// TIA Portal project "Delta_Praktika_P&P" (V17) (continued)

               // jog to position
               //*********************************************************************************************************
             ELSIF #tempJogToPosition THEN
               // set jog target position and configuration
               #instMC_MoveLinearAbsoute.Position[1] := #targetPosition.x;
               #instMC_MoveLinearAbsoute.Position[2] := #targetPosition.y;
               #instMC_MoveLinearAbsoute.Position[3] := #targetPosition.z;
               #instMC_MoveLinearAbsoute.Position[4] := #targetPosition.a;
               #instMC_MoveLinearAbsoute.CoordSystem := #coordSystem;
               #instMC_MoveLinearAbsoute.Velocity := #dynamics.path.velocity;
               #instMC_MoveLinearAbsoute.Acceleration := #dynamics.path.acceleration;
               #instMC_MoveLinearAbsoute.Deceleration := #dynamics.path.deceleration;
               #instMC_MoveLinearAbsoute.Jerk := #dynamics.path.jerk;
               #instMC_MoveLinearAbsoute.DynamicAdaption := #dynamics.dynamicAdaption;
               #instMC_MoveLinearAbsoute.DirectionA := #dynamics.directionA;

               // jog synchronous point to point
               //*********************************************************************************************************
             ELSIF #tempJogSPTP THEN
               #instMC_MoveDirectAbsolute.Position[1] := #targetPosition.x;
               #instMC_MoveDirectAbsolute.Position[2] := #targetPosition.y;
               #instMC_MoveDirectAbsolute.Position[3] := #targetPosition.z;
               #instMC_MoveDirectAbsolute.Position[4] := #targetPosition.a;
               #instMC_MoveDirectAbsolute.CoordSystem := #coordSystem;
               #instMC_MoveDirectAbsolute.VelocityFactor := #dynamics.sPTP.velocityFactor;
               #instMC_MoveDirectAbsolute.AccelerationFactor := #dynamics.sPTP.accelerationFactor;
               #instMC_MoveDirectAbsolute.DecelerationFactor := #dynamics.sPTP.decelerationFactor;
               #instMC_MoveDirectAbsolute.JerkFactor := #dynamics.sPTP.jerkFactor;
               #instMC_MoveDirectAbsolute.LinkConstellation := #linkconstellation;
               #instMC_MoveDirectAbsolute.PositionMode := 1;
               #instMC_MoveDirectAbsolute.DirectionA := #dynamics.directionA;

             END_IF;

           END_REGION

           REGION SET_ORIENTATION_DYNAMICS

             IF (((#jogDirection = 4) AND (#tempJogForward OR #tempJogBackward)) OR #tempJogToPosition)
               AND (#dynamics.orientation.velocity > 0.0 // check if change of orientation dynamics is required
               OR #dynamics.orientation.acceleration > 0.0
               OR #dynamics.orientation.deceleration > 0.0
               OR #dynamics.orientation.jerk > 0.0)
             THEN
               // safe default dynamics for orientation axis
               #statOrientationDynamicsOld.velocity := #axesGroup.DynamicDefaults.Orientation.Velocity;
               #statOrientationDynamicsOld.acceleration := #axesGroup.DynamicDefaults.Orientation.Acceleration;
               #statOrientationDynamicsOld.deceleration := #axesGroup.DynamicDefaults.Orientation.Deceleration;
               #statOrientationDynamicsOld.jerk := #axesGroup.DynamicDefaults.Orientation.Jerk;

               // change orientation default dynamics temporary
               IF #dynamics.orientation.velocity > 0.0 THEN
                 #axesGroup.DynamicDefaults.Orientation.Velocity := #dynamics.orientation.velocity;
               END_IF;
               IF #dynamics.orientation.acceleration > 0.0 THEN
                 #axesGroup.DynamicDefaults.Orientation.Acceleration := #dynamics.orientation.acceleration;
               END_IF;
               IF #dynamics.orientation.deceleration > 0.0 THEN
                 #axesGroup.DynamicDefaults.Orientation.Deceleration := #dynamics.orientation.deceleration;
               END_IF;
               IF #dynamics.orientation.jerk > 0.0 THEN
                 #axesGroup.DynamicDefaults.Orientation.Jerk := #dynamics.orientation.jerk;
               END_IF;

               // Orientation default dynamics will be reseted to previous values after jogging
               #statOrientationDynamicsChanged := TRUE;
             END_IF;
           END_REGION

           REGION STATE_TRANSITION

             // check if change of tool is required
             IF (#tool <> #statToolOld) THEN
               #statFBState := #FB_STATE_SET_TOOL;
             ELSE // execute movement
               #statFBState := #FB_STATE_EXECUTE_MOVEMENT;
             END_IF;

           END_REGION

         END_IF;

       #FB_STATE_SET_TOOL:

         REGION TOOL_CHANGE

           IF #axesGroup.StatusWord.%X6 // no motion command is acitve
             AND NOT #axesGroup.StatusWord.%X17 // not interrupted
             AND #axesGroup.StatusWord.%X12 // constant velocity
           THEN
             #instMC_SetTool.Execute := TRUE;
             #instMC_SetTool.ToolNumber := #tool;
           END_IF;

         END_REGION

         REGION STATE_TRANSITION

           // tool has been changed
           IF #instMC_SetTool.Done THEN
             #statToolOld := #tool;
             #statFBState := #FB_STATE_EXECUTE_MOVEMENT;
           END_IF;

         END_REGION

       #FB_STATE_EXECUTE_MOVEMENT:

         REGION SET_JOG_COMMAND

             // Cartesian jogging
             IF (#tempJogForward OR #tempJogBackward) THEN
               #instMC_MoveLinearRelative.Execute := TRUE;

               // jog to target position  
             ELSIF #tempJogToPosition THEN
               #instMC_MoveLinearAbsoute.Execute := TRUE;

               //jog synchronous point to point
             ELSIF #tempJogSPTP THEN
               #instMC_MoveDirectAbsolute.Execute := TRUE;

             ELSE
               #instMC_MoveLinearRelative.Execute := FALSE;
               #instMC_MoveLinearAbsoute.Execute := FALSE;
               #instMC_MoveDirectAbsolute.Execute := FALSE;
             END_IF;

         END_REGION

         REGION STATE_TRANSITION

           IF #instMC_MoveLinearRelative.Done OR #instMC_MoveLinearAbsoute.Done OR #instMC_MoveDirectAbsolute.Done THEN
             #statStatus := #STATUS_EXECUTION_FINISHED;
           END_IF;

         END_REGION

       #FB_STATE_STOP:

         REGION STOP_KINEMATICS_MOTION

           // set execute if group stop not busy
           #instMC_GroupStop.Execute := (NOT #instMC_GroupStop.Busy AND NOT #instMC_GroupStop.Done AND NOT #instMC_GroupStop.Error);

         END_REGION

         REGION STATE_TRANSITION

           IF (#instMC_GroupStop.Done AND #axesGroup.StatusWord.%X6) THEN // Added X6 according to AW
             #statStatus := #STATUS_EXECUTION_FINISHED;
           ELSIF #axesGroup.StatusWord.%X1 THEN // general TO error
             #statStatus := #ERR_TO_KINEMATICS;
           ELSIF #instMC_MoveLinearRelative.Error THEN
             #statStatus := #instMC_MoveLinearRelative.ErrorId;
           ELSIF #instMC_MoveLinearAbsoute.Error THEN
             #statStatus := #instMC_MoveLinearAbsoute.ErrorId;
           ELSIF #instMC_MoveDirectAbsolute.Error THEN
             #statStatus := #instMC_MoveDirectAbsolute.ErrorId;
           ELSIF #instMC_SetTool.Error THEN
             #statStatus := #instMC_SetTool.ErrorId;
           ELSIF #instMC_GroupStop.Error THEN
             #statStatus := #instMC_GroupStop.ErrorId;
           END_IF;

         END_REGION

       ELSE // Undefined state in state machine reached
         #statStatus := #ERR_UNDEFINED_STATE;
     END_CASE;

   END_REGION STATE_MACHINE

   REGION OUTPUTS

     // Write outputs
     IF (#statStatus = #STATUS_EXECUTION_FINISHED) AND (#statDone = FALSE) AND (#statError = FALSE) THEN // Execution finished without errors
       #statDone := TRUE;
       #statBusy := FALSE;
       #statActive := FALSE;
       #statError := FALSE;
       #statFBState := #FB_STATE_NO_PROCESSING; // Switch state machine to "no processing"

     ELSIF (#statStatus.%X15 = TRUE) AND (#statError = FALSE) THEN // Error occurred (#statStatus is 16#8000 to 16#FFFF)
       #statDone := FALSE;
       #statBusy := FALSE;
       #statActive := FALSE;
       #statError := TRUE;
       // Write diagnostics
       #tempRet := RD_SYS_T(#diagnostics.timeStamp);
       #diagnostics.stateNumber := #statFBState;
       #diagnostics.status := #statStatus;
       #statFBState := #FB_STATE_NO_PROCESSING; // Switch state machine to "no processing"

     ELSIF (#tempJogForward = FALSE AND #tempJogBackward = FALSE AND #tempJogToPosition = FALSE AND #tempJogSPTP = FALSE) AND ((#statDone = TRUE) OR (#statError = TRUE)) THEN // Reset outputs
       #statDone := FALSE;
       #statBusy := FALSE;
       #statActive := FALSE;
       #statError := FALSE;
       #statStatus := #STATUS_NO_CALL;
       #statJogForwardOld := FALSE;
       #statJogBackwardOld := FALSE;
       #statJogToPositionOld := FALSE;
       #statJogSPTPOld := FALSE;
     END_IF;

     // Write static values to outputs
     #done := #statDone;
     #busy := #statBusy;
     #active := #statActive;
     #error := #statError;
     #status := #statStatus;
     #remainingDistance := #statRemainingDistance;

   END_REGION OUTPUTS

   REGION CALL_FB_CYCLICALLY

     // call FBs and set Execute = FALSE after the call
     #instMC_GroupStop(AxesGroup := #axesGroup);
     #instMC_GroupStop.Execute := FALSE;

     #instMC_MoveLinearAbsoute(AxesGroup := #axesGroup);
     #instMC_MoveLinearAbsoute.Execute := FALSE;

     #instMC_MoveLinearRelative(AxesGroup := #axesGroup);
     #instMC_MoveLinearRelative.Execute := FALSE;

     #instMC_SetTool(AxesGroup := #axesGroup);
     #instMC_SetTool.Execute := FALSE;

     #instMC_MoveDirectAbsolute(AxesGroup := #axesGroup);
     #instMC_MoveDirectAbsolute.Execute := FALSE;
   END_REGION
END_FUNCTION_BLOCK

FUNCTION "Sekuentzia" : Void   // FC1, LAD
{ S7_Optimized_Access := 'TRUE' }
VERSION : 0.1
   VAR_TEMP   // added for the SCL form of the ladder/FBD networks
      _w1 : Bool;
   END_VAR
BEGIN

REGION Network 1
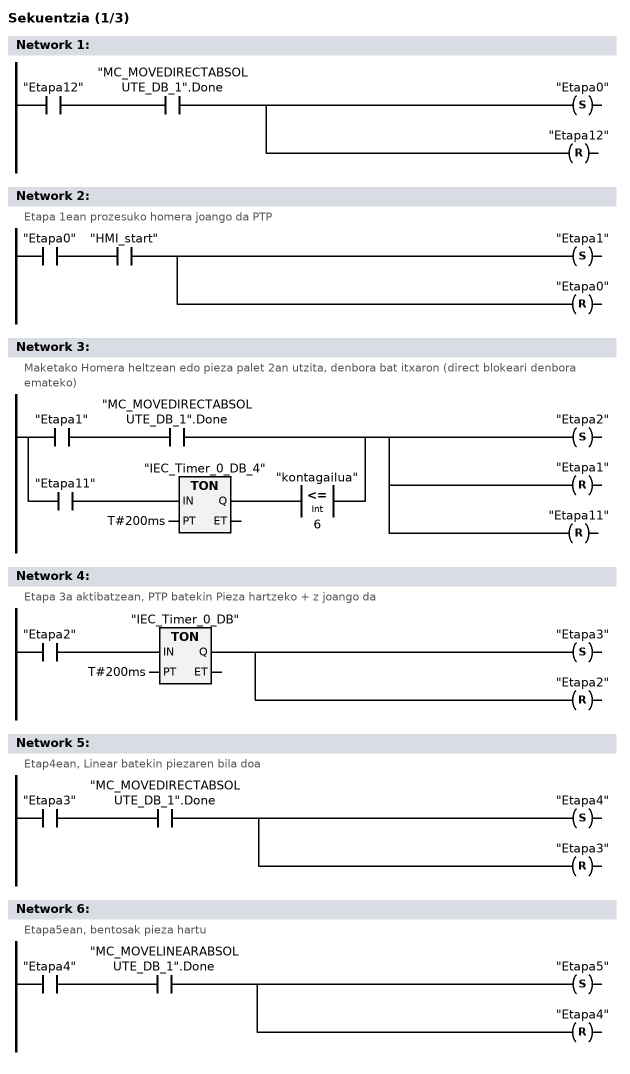
   RUNG wire#powerrail
      Contact( "Etapa12" )
      Contact( "MC_MOVEDIRECTABSOLUTE_DB_1".Done )
      wire#w1
      S_Coil( "Etapa0" )
   END_RUNG
   RUNG wire#w1
      R_Coil( "Etapa12" )
   END_RUNG
   // the same network as SCL:
   IF "Etapa12" AND "MC_MOVEDIRECTABSOLUTE_DB_1".Done THEN
       "Etapa0" := TRUE;
       "Etapa12" := FALSE;
   END_IF;
END_REGION

REGION Network 2
   // Etapa 1ean prozesuko homera joango da PTP
   RUNG wire#powerrail
      Contact( "Etapa0" )
      Contact( "HMI_start" )
      wire#w1
      S_Coil( "Etapa1" )
   END_RUNG
   RUNG wire#w1
      R_Coil( "Etapa0" )
   END_RUNG
   // the same network as SCL:
   IF "Etapa0" AND "HMI_start" THEN
       "Etapa1" := TRUE;
       "Etapa0" := FALSE;
   END_IF;
END_REGION

REGION Network 3
   // Maketako Homera heltzean edo pieza palet 2an utzita, denbora bat itxaron (direct blokeari denbora emateko)
   "IEC_Timer_0_DB_4".TON(IN := "Etapa11", PT := T#200ms);
   IF ("Etapa1" AND "MC_MOVEDIRECTABSOLUTE_DB_1".Done) OR ("IEC_Timer_0_DB_4".Q AND ("kontagailua" <= 6)) THEN
       "Etapa2" := TRUE;
   END_IF;
   #_w1 := ("Etapa1" AND "MC_MOVEDIRECTABSOLUTE_DB_1".Done) OR ("IEC_Timer_0_DB_4".Q AND ("kontagailua" <= 6));
   IF #_w1 THEN
       "Etapa1" := FALSE;
       "Etapa11" := FALSE;
   END_IF;
END_REGION

REGION Network 4
   // Etapa 3a aktibatzean, PTP batekin Pieza hartzeko + z joango da
   "IEC_Timer_0_DB".TON(IN := "Etapa2", PT := T#200ms);
   IF "IEC_Timer_0_DB".Q THEN
       "Etapa3" := TRUE;
       "Etapa2" := FALSE;
   END_IF;
END_REGION

REGION Network 5
   // Etap4ean, Linear batekin piezaren bila doa
   RUNG wire#powerrail
      Contact( "Etapa3" )
      Contact( "MC_MOVEDIRECTABSOLUTE_DB_1".Done )
      wire#w1
      S_Coil( "Etapa4" )
   END_RUNG
   RUNG wire#w1
      R_Coil( "Etapa3" )
   END_RUNG
   // the same network as SCL:
   IF "Etapa3" AND "MC_MOVEDIRECTABSOLUTE_DB_1".Done THEN
       "Etapa4" := TRUE;
       "Etapa3" := FALSE;
   END_IF;
END_REGION

REGION Network 6
   // Etapa5ean, bentosak pieza hartu
   RUNG wire#powerrail
      Contact( "Etapa4" )
      Contact( "MC_MOVELINEARABSOLUTE_DB_1".Done )
      wire#w1
      S_Coil( "Etapa5" )
   END_RUNG
   RUNG wire#w1
      R_Coil( "Etapa4" )
   END_RUNG
   // the same network as SCL:
   IF "Etapa4" AND "MC_MOVELINEARABSOLUTE_DB_1".Done THEN
       "Etapa5" := TRUE;
       "Etapa4" := FALSE;
   END_IF;
END_REGION

REGION Network 7
   // Denbora bat eman eta etapa6an Linear batekin z+
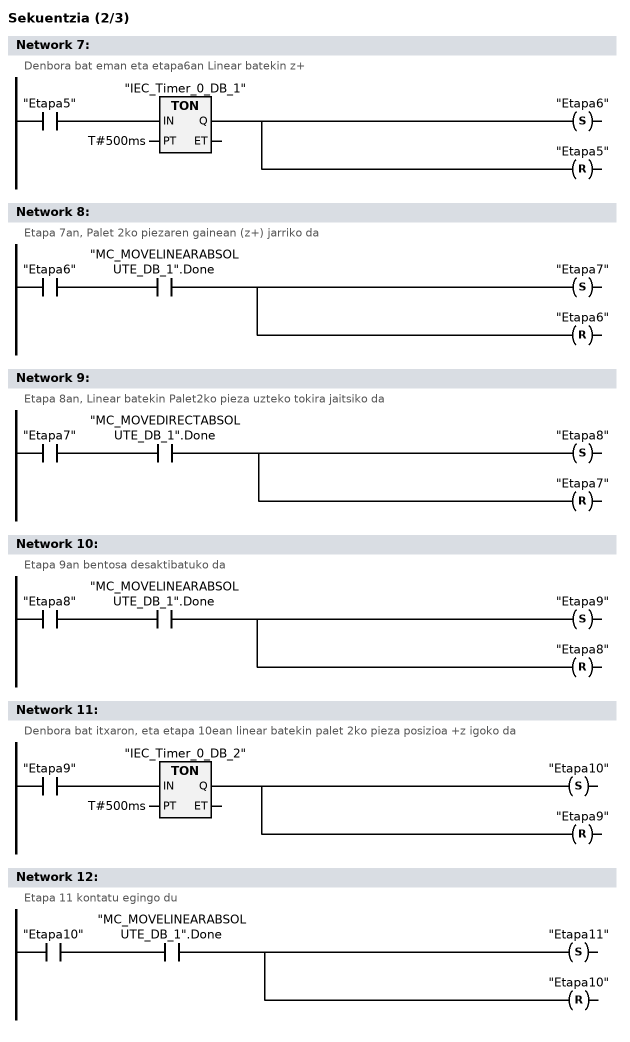
   "IEC_Timer_0_DB_1".TON(IN := "Etapa5", PT := T#500ms);
   IF "IEC_Timer_0_DB_1".Q THEN
       "Etapa6" := TRUE;
       "Etapa5" := FALSE;
   END_IF;
END_REGION

REGION Network 8
   // Etapa 7an, Palet 2ko piezaren gainean (z+) jarriko da
   RUNG wire#powerrail
      Contact( "Etapa6" )
      Contact( "MC_MOVELINEARABSOLUTE_DB_1".Done )
      wire#w1
      S_Coil( "Etapa7" )
   END_RUNG
   RUNG wire#w1
      R_Coil( "Etapa6" )
   END_RUNG
   // the same network as SCL:
   IF "Etapa6" AND "MC_MOVELINEARABSOLUTE_DB_1".Done THEN
       "Etapa7" := TRUE;
       "Etapa6" := FALSE;
   END_IF;
END_REGION

REGION Network 9
   // Etapa 8an, Linear batekin Palet2ko pieza uzteko tokira jaitsiko da
   RUNG wire#powerrail
      Contact( "Etapa7" )
      Contact( "MC_MOVEDIRECTABSOLUTE_DB_1".Done )
      wire#w1
      S_Coil( "Etapa8" )
   END_RUNG
   RUNG wire#w1
      R_Coil( "Etapa7" )
   END_RUNG
   // the same network as SCL:
   IF "Etapa7" AND "MC_MOVEDIRECTABSOLUTE_DB_1".Done THEN
       "Etapa8" := TRUE;
       "Etapa7" := FALSE;
   END_IF;
END_REGION

REGION Network 10
   // Etapa 9an bentosa desaktibatuko da
   RUNG wire#powerrail
      Contact( "Etapa8" )
      Contact( "MC_MOVELINEARABSOLUTE_DB_1".Done )
      wire#w1
      S_Coil( "Etapa9" )
   END_RUNG
   RUNG wire#w1
      R_Coil( "Etapa8" )
   END_RUNG
   // the same network as SCL:
   IF "Etapa8" AND "MC_MOVELINEARABSOLUTE_DB_1".Done THEN
       "Etapa9" := TRUE;
       "Etapa8" := FALSE;
   END_IF;
END_REGION

REGION Network 11
   // Denbora bat itxaron, eta etapa 10ean linear batekin palet 2ko pieza posizioa +z igoko da
   "IEC_Timer_0_DB_2".TON(IN := "Etapa9", PT := T#500ms);
   IF "IEC_Timer_0_DB_2".Q THEN
       "Etapa10" := TRUE;
       "Etapa9" := FALSE;
   END_IF;
END_REGION

REGION Network 12
   // Etapa 11 kontatu egingo du
   RUNG wire#powerrail
      Contact( "Etapa10" )
      Contact( "MC_MOVELINEARABSOLUTE_DB_1".Done )
      wire#w1
      S_Coil( "Etapa11" )
   END_RUNG
   RUNG wire#w1
      R_Coil( "Etapa10" )
   END_RUNG
   // the same network as SCL:
   IF "Etapa10" AND "MC_MOVELINEARABSOLUTE_DB_1".Done THEN
       "Etapa11" := TRUE;
       "Etapa10" := FALSE;
   END_IF;
END_REGION

REGION Network 13
   // Etapa 11 + denbora bat pasatzean, zenbat kontatu dituen ikusten du 6 baino gehiago bada, etapa 12an PTP batekin maketaren homera joango da
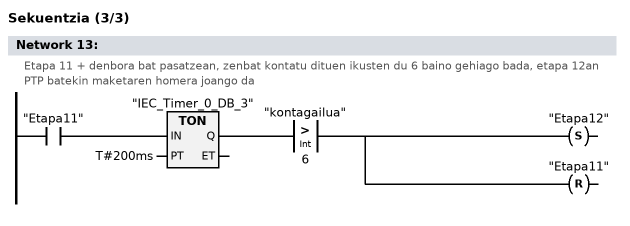
   "IEC_Timer_0_DB_3".TON(IN := "Etapa11", PT := T#200ms);
   IF "IEC_Timer_0_DB_3".Q AND ("kontagailua" > 6) THEN
       "Etapa12" := TRUE;
       "Etapa11" := FALSE;
   END_IF;
END_REGION
END_FUNCTION

FUNCTION "Mugimeduak" : Void   // FC2, LAD
{ S7_Optimized_Access := 'TRUE' }
VERSION : 0.1
BEGIN

REGION Network 1
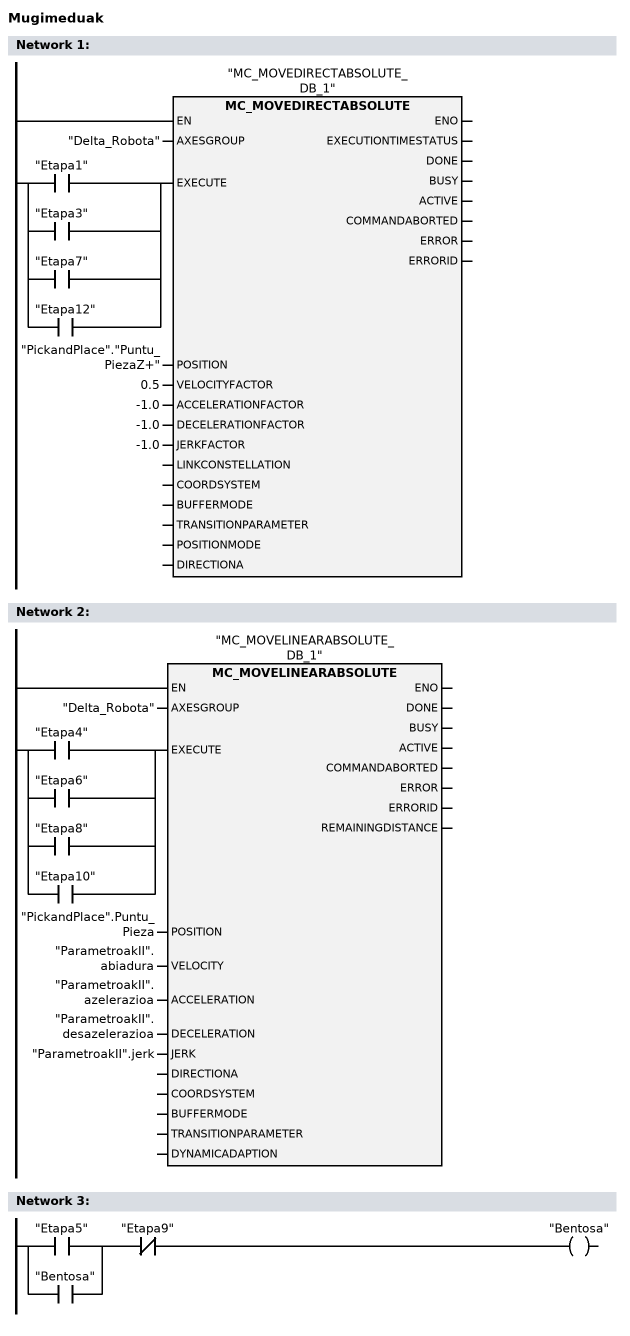
   "MC_MOVEDIRECTABSOLUTE_DB_1"(AxesGroup := "Delta_Robota",   // MC_MOVEDIRECTABSOLUTE
                           Execute := "Etapa1" OR "Etapa3" OR "Etapa7" OR "Etapa12",
                           Position := "PickandPlace"."Puntu_PiezaZ+",
                           VelocityFactor := 0.5,
                           AccelerationFactor := -1.0,
                           DecelerationFactor := -1.0,
                           JerkFactor := -1.0);
END_REGION

REGION Network 2
   "MC_MOVELINEARABSOLUTE_DB_1"(AxesGroup := "Delta_Robota",   // MC_MOVELINEARABSOLUTE
                           Execute := "Etapa4" OR "Etapa6" OR "Etapa8" OR "Etapa10",
                           Position := "PickandPlace".Puntu_Pieza,
                           Velocity := "ParametroakII".abiadura,
                           Acceleration := "ParametroakII".azelerazioa,
                           Deceleration := "ParametroakII".desazelerazioa,
                           Jerk := "ParametroakII".jerk);
END_REGION

REGION Network 3
   RUNG wire#powerrail
      Contact( "Etapa5" )
      wire#w1
      I_Contact( "Etapa9" )
      Coil( "Bentosa" )
   END_RUNG
   RUNG wire#powerrail
      Contact( "Bentosa" )
   END_RUNG wire#w1
   // the same network as SCL:
   "Bentosa" := ("Etapa5" OR "Bentosa") AND NOT "Etapa9";
END_REGION
END_FUNCTION

FUNCTION "Kontagailu_sek" : Void   // FC3, LAD
{ S7_Optimized_Access := 'TRUE' }
VERSION : 0.1
   VAR_TEMP   // added for the SCL form of the ladder/FBD networks
      _w1 : Bool;
      _w2 : Bool;
      _w3 : Bool;
   END_VAR
BEGIN

REGION Network 1
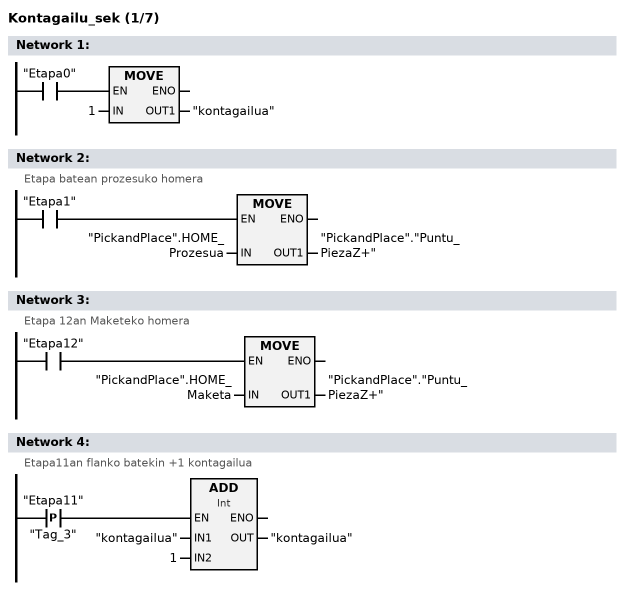
   RUNG wire#powerrail
      Contact( "Etapa0" )
      Move(in := 1, out1 => "kontagailua")
   END_RUNG
   // the same network as SCL:
   IF "Etapa0" THEN "kontagailua" := 1; END_IF;
END_REGION

REGION Network 2
   // Etapa batean prozesuko homera
   RUNG wire#powerrail
      Contact( "Etapa1" )
      Move(in := "PickandPlace".HOME_Prozesua, out1 => "PickandPlace"."Puntu_PiezaZ+")
   END_RUNG
   // the same network as SCL:
   IF "Etapa1" THEN "PickandPlace"."Puntu_PiezaZ+" := "PickandPlace".HOME_Prozesua; END_IF;
END_REGION

REGION Network 3
   // Etapa 12an Maketeko homera
   RUNG wire#powerrail
      Contact( "Etapa12" )
      Move(in := "PickandPlace".HOME_Maketa, out1 => "PickandPlace"."Puntu_PiezaZ+")
   END_RUNG
   // the same network as SCL:
   IF "Etapa12" THEN "PickandPlace"."Puntu_PiezaZ+" := "PickandPlace".HOME_Maketa; END_IF;
END_REGION

REGION Network 4
   // Etapa11an flanko batekin +1 kontagailua
   RUNG wire#powerrail
      P_Contact(operand := "Etapa11", bit := "Tag_3")
      { S7_Templates := "SrcType := Int" } Add(in1 := "kontagailua", in2 := 1, out => "kontagailua")
   END_RUNG
   // the same network as SCL:
   #_w1 := "Etapa11" AND NOT "Tag_3";   // rising edge of "Etapa11"
   "Tag_3" := "Etapa11";
   IF #_w1 THEN "kontagailua" := "kontagailua" + 1; END_IF;
END_REGION

REGION Network 5
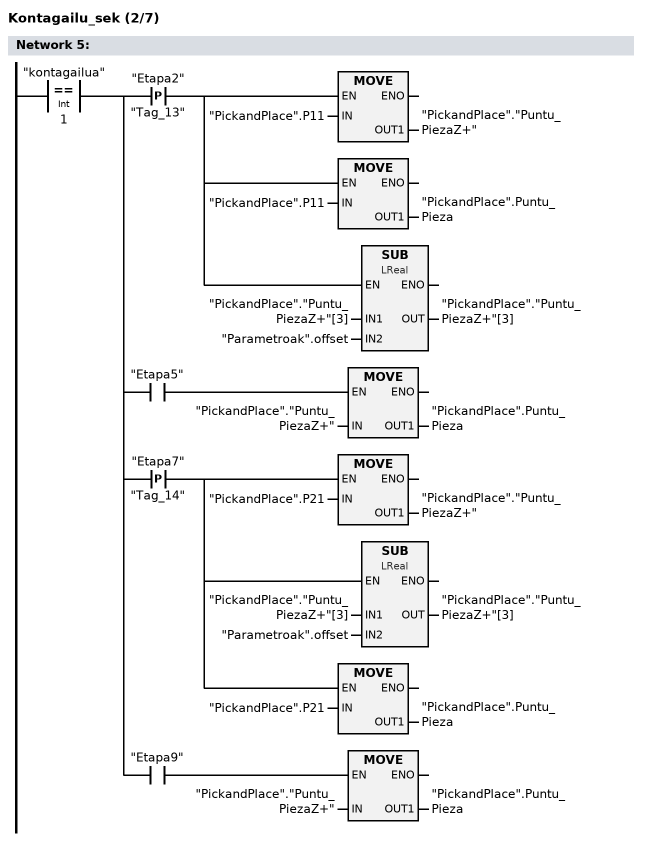
   RUNG wire#powerrail
      { S7_Templates := "SrcType := Int" } EQ_Contact(in1 := "kontagailua", in2 := 1)
      wire#w1
      P_Contact(operand := "Etapa2", bit := "Tag_13")
      wire#w2
      Move(in := "PickandPlace".P11, out1 => "PickandPlace"."Puntu_PiezaZ+")
   END_RUNG
   RUNG wire#w2
      Move(in := "PickandPlace".P11, out1 => "PickandPlace".Puntu_Pieza)
   END_RUNG
   RUNG wire#w2
      { S7_Templates := "SrcType := LReal" } Sub(in1 := "PickandPlace"."Puntu_PiezaZ+"[3], in2 := "Parametroak".offset, out => "PickandPlace"."Puntu_PiezaZ+"[3])
   END_RUNG
   RUNG wire#w1
      Contact( "Etapa5" )
      Move(in := "PickandPlace"."Puntu_PiezaZ+", out1 => "PickandPlace".Puntu_Pieza)
   END_RUNG
   RUNG wire#w1
      P_Contact(operand := "Etapa7", bit := "Tag_14")
      wire#w3
      Move(in := "PickandPlace".P21, out1 => "PickandPlace"."Puntu_PiezaZ+")
   END_RUNG
   RUNG wire#w3
      { S7_Templates := "SrcType := LReal" } Sub(in1 := "PickandPlace"."Puntu_PiezaZ+"[3], in2 := "Parametroak".offset, out => "PickandPlace"."Puntu_PiezaZ+"[3])
   END_RUNG
   RUNG wire#w3
      Move(in := "PickandPlace".P21, out1 => "PickandPlace".Puntu_Pieza)
   END_RUNG
   RUNG wire#w1
      Contact( "Etapa9" )
      Move(in := "PickandPlace"."Puntu_PiezaZ+", out1 => "PickandPlace".Puntu_Pieza)
   END_RUNG
   // the same network as SCL:
   #_w1 := "kontagailua" = 1;
   #_w2 := #_w1 AND "Etapa2" AND NOT "Tag_13";   // rising edge of "Etapa2"
   "Tag_13" := "Etapa2";
   IF #_w2 THEN
       "PickandPlace"."Puntu_PiezaZ+" := "PickandPlace".P11;
       "PickandPlace".Puntu_Pieza := "PickandPlace".P11;
       "PickandPlace"."Puntu_PiezaZ+"[3] := "PickandPlace"."Puntu_PiezaZ+"[3] - "Parametroak".offset;
   END_IF;
   IF #_w1 AND "Etapa5" THEN "PickandPlace".Puntu_Pieza := "PickandPlace"."Puntu_PiezaZ+"; END_IF;
   #_w3 := #_w1 AND "Etapa7" AND NOT "Tag_14";   // rising edge of "Etapa7"
   "Tag_14" := "Etapa7";
   IF #_w3 THEN
       "PickandPlace"."Puntu_PiezaZ+" := "PickandPlace".P21;
       "PickandPlace"."Puntu_PiezaZ+"[3] := "PickandPlace"."Puntu_PiezaZ+"[3] - "Parametroak".offset;
       "PickandPlace".Puntu_Pieza := "PickandPlace".P21;
   END_IF;
   IF #_w1 AND "Etapa9" THEN "PickandPlace".Puntu_Pieza := "PickandPlace"."Puntu_PiezaZ+"; END_IF;
END_REGION

REGION Network 6
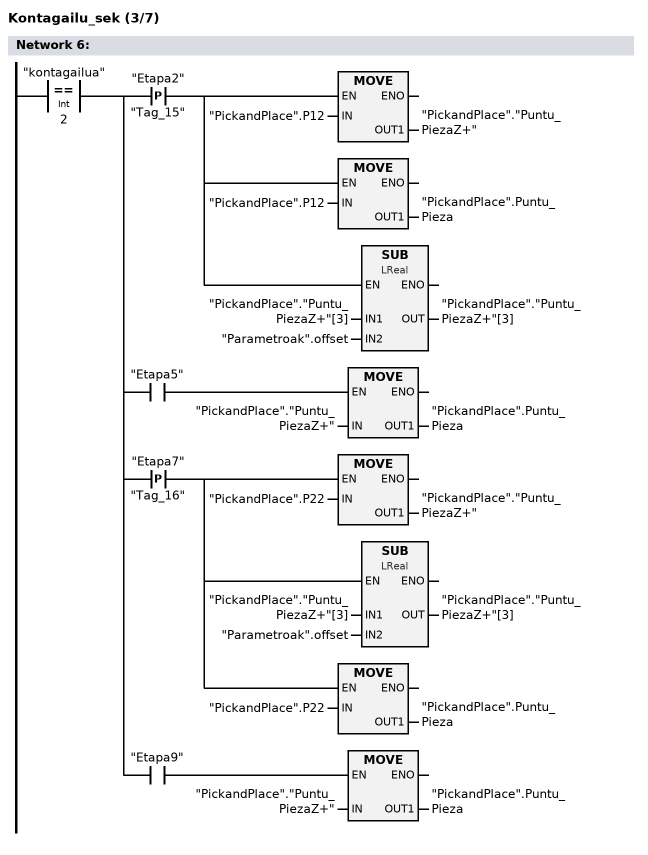
   RUNG wire#powerrail
      { S7_Templates := "SrcType := Int" } EQ_Contact(in1 := "kontagailua", in2 := 2)
      wire#w1
      P_Contact(operand := "Etapa2", bit := "Tag_15")
      wire#w2
      Move(in := "PickandPlace".P12, out1 => "PickandPlace"."Puntu_PiezaZ+")
   END_RUNG
   RUNG wire#w2
      Move(in := "PickandPlace".P12, out1 => "PickandPlace".Puntu_Pieza)
   END_RUNG
   RUNG wire#w2
      { S7_Templates := "SrcType := LReal" } Sub(in1 := "PickandPlace"."Puntu_PiezaZ+"[3], in2 := "Parametroak".offset, out => "PickandPlace"."Puntu_PiezaZ+"[3])
   END_RUNG
   RUNG wire#w1
      Contact( "Etapa5" )
      Move(in := "PickandPlace"."Puntu_PiezaZ+", out1 => "PickandPlace".Puntu_Pieza)
   END_RUNG
   RUNG wire#w1
      P_Contact(operand := "Etapa7", bit := "Tag_16")
      wire#w3
      Move(in := "PickandPlace".P22, out1 => "PickandPlace"."Puntu_PiezaZ+")
   END_RUNG
   RUNG wire#w3
      { S7_Templates := "SrcType := LReal" } Sub(in1 := "PickandPlace"."Puntu_PiezaZ+"[3], in2 := "Parametroak".offset, out => "PickandPlace"."Puntu_PiezaZ+"[3])
   END_RUNG
   RUNG wire#w3
      Move(in := "PickandPlace".P22, out1 => "PickandPlace".Puntu_Pieza)
   END_RUNG
   RUNG wire#w1
      Contact( "Etapa9" )
      Move(in := "PickandPlace"."Puntu_PiezaZ+", out1 => "PickandPlace".Puntu_Pieza)
   END_RUNG
   // the same network as SCL:
   #_w1 := "kontagailua" = 2;
   #_w2 := #_w1 AND "Etapa2" AND NOT "Tag_15";   // rising edge of "Etapa2"
   "Tag_15" := "Etapa2";
   IF #_w2 THEN
       "PickandPlace"."Puntu_PiezaZ+" := "PickandPlace".P12;
       "PickandPlace".Puntu_Pieza := "PickandPlace".P12;
       "PickandPlace"."Puntu_PiezaZ+"[3] := "PickandPlace"."Puntu_PiezaZ+"[3] - "Parametroak".offset;
   END_IF;
   IF #_w1 AND "Etapa5" THEN "PickandPlace".Puntu_Pieza := "PickandPlace"."Puntu_PiezaZ+"; END_IF;
   #_w3 := #_w1 AND "Etapa7" AND NOT "Tag_16";   // rising edge of "Etapa7"
   "Tag_16" := "Etapa7";
   IF #_w3 THEN
       "PickandPlace"."Puntu_PiezaZ+" := "PickandPlace".P22;
       "PickandPlace"."Puntu_PiezaZ+"[3] := "PickandPlace"."Puntu_PiezaZ+"[3] - "Parametroak".offset;
       "PickandPlace".Puntu_Pieza := "PickandPlace".P22;
   END_IF;
   IF #_w1 AND "Etapa9" THEN "PickandPlace".Puntu_Pieza := "PickandPlace"."Puntu_PiezaZ+"; END_IF;
END_REGION

REGION Network 7
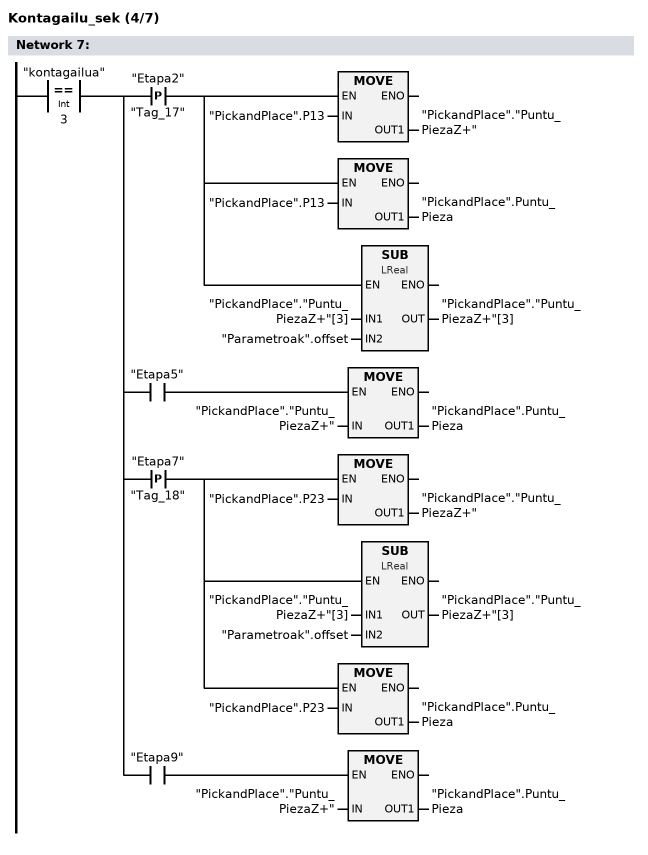
   RUNG wire#powerrail
      { S7_Templates := "SrcType := Int" } EQ_Contact(in1 := "kontagailua", in2 := 3)
      wire#w1
      P_Contact(operand := "Etapa2", bit := "Tag_17")
      wire#w2
      Move(in := "PickandPlace".P13, out1 => "PickandPlace"."Puntu_PiezaZ+")
   END_RUNG
   RUNG wire#w2
      Move(in := "PickandPlace".P13, out1 => "PickandPlace".Puntu_Pieza)
   END_RUNG
   RUNG wire#w2
      { S7_Templates := "SrcType := LReal" } Sub(in1 := "PickandPlace"."Puntu_PiezaZ+"[3], in2 := "Parametroak".offset, out => "PickandPlace"."Puntu_PiezaZ+"[3])
   END_RUNG
   RUNG wire#w1
      Contact( "Etapa5" )
      Move(in := "PickandPlace"."Puntu_PiezaZ+", out1 => "PickandPlace".Puntu_Pieza)
   END_RUNG
   RUNG wire#w1
      P_Contact(operand := "Etapa7", bit := "Tag_18")
      wire#w3
      Move(in := "PickandPlace".P23, out1 => "PickandPlace"."Puntu_PiezaZ+")
   END_RUNG
   RUNG wire#w3
      { S7_Templates := "SrcType := LReal" } Sub(in1 := "PickandPlace"."Puntu_PiezaZ+"[3], in2 := "Parametroak".offset, out => "PickandPlace"."Puntu_PiezaZ+"[3])
   END_RUNG
   RUNG wire#w3
      Move(in := "PickandPlace".P23, out1 => "PickandPlace".Puntu_Pieza)
   END_RUNG
   RUNG wire#w1
      Contact( "Etapa9" )
      Move(in := "PickandPlace"."Puntu_PiezaZ+", out1 => "PickandPlace".Puntu_Pieza)
   END_RUNG
   // the same network as SCL:
   #_w1 := "kontagailua" = 3;
   #_w2 := #_w1 AND "Etapa2" AND NOT "Tag_17";   // rising edge of "Etapa2"
   "Tag_17" := "Etapa2";
   IF #_w2 THEN
       "PickandPlace"."Puntu_PiezaZ+" := "PickandPlace".P13;
       "PickandPlace".Puntu_Pieza := "PickandPlace".P13;
       "PickandPlace"."Puntu_PiezaZ+"[3] := "PickandPlace"."Puntu_PiezaZ+"[3] - "Parametroak".offset;
   END_IF;
   IF #_w1 AND "Etapa5" THEN "PickandPlace".Puntu_Pieza := "PickandPlace"."Puntu_PiezaZ+"; END_IF;
   #_w3 := #_w1 AND "Etapa7" AND NOT "Tag_18";   // rising edge of "Etapa7"
   "Tag_18" := "Etapa7";
   IF #_w3 THEN
       "PickandPlace"."Puntu_PiezaZ+" := "PickandPlace".P23;
       "PickandPlace"."Puntu_PiezaZ+"[3] := "PickandPlace"."Puntu_PiezaZ+"[3] - "Parametroak".offset;
       "PickandPlace".Puntu_Pieza := "PickandPlace".P23;
   END_IF;
   IF #_w1 AND "Etapa9" THEN "PickandPlace".Puntu_Pieza := "PickandPlace"."Puntu_PiezaZ+"; END_IF;
END_REGION

REGION Network 8